(* Logix 5000 project; controller PLC_MCC1300_75F1 vendor 1 type 14 code 166 rev 32.11; software revision 32.04; part 18 of 83 *)
(* tags used below, declared in another part *)
   GP_OB_InitializeMain : GP_OB_Initialize;
   M302SpeedUp : MAC_SpeedUp;
   M310_M4_DR_B1 : AXIS_CIP_DRIVE;
   M310B : MAC_Conveyor;
   M310B_ALM : MAC_Conveyor_ALM;
   M310B_Data : UDT_Convoy_SL;
   M310B_HMR : MAC_Conveyor_HMR;
   M310B_HMW : MAC_Conveyor_HMW;
   M310B_M1_DR_IN_MAJ : MOTION_INSTRUCTION;
   M310B_M1_DR_IN_MAR : MOTION_INSTRUCTION;
   M310B_M1_DR_IN_MAS : MOTION_INSTRUCTION;
   M310B_M1_DR_IN_MRP : MOTION_INSTRUCTION;
   M310B_M1_DR_MAFR : MOTION_INSTRUCTION;
   M310B_M1_DR_MDR : MOTION_INSTRUCTION;
   M310B_M1_DR_MSF : MOTION_INSTRUCTION;
   M310B_M1_DR_MSO : MOTION_INSTRUCTION;
   M310B_M1_DR_OUT_MAJ : MOTION_INSTRUCTION;
   M310B_M1_DR_OUT_MAM : MOTION_INSTRUCTION;
   M310B_M1_DR_OUT_MAR : MOTION_INSTRUCTION;
   M310B_M1_DR_OUT_MCD : MOTION_INSTRUCTION;
   M310B_M1_DR_OUT_MRP : MOTION_INSTRUCTION;
   M310B_SpaceConv_Utilities : SpaceConv_Utilities;
   M310B_xOS_PosReq : BOOL;
   M311 : MAC_Conveyor;
   TMP_d : DINT;
   TMP_dDirection : DINT;
   TMP_r : REAL;
   TMP_rAcc : REAL;
   TMP_rDec : REAL;
   TMP_rSpeed : REAL;
   TMP_rTarget_M1 : REAL;
   TMP_xForwardCommadnForCleaningZone : BOOL;
   TMP_xPositioning : BOOL;
   TMP_xPositioning_M1 : BOOL;
   TMP_xPositioning_M2 : BOOL;
   TMP_xPowerSaving : BOOL;
   TMP_xReverse : BOOL;
   TMP_xReverse_M1 : BOOL;
   TMP_xReverse_M2 : BOOL;
   TMP_xRun : BOOL;
   TMP_xRun_M1 : BOOL;
   TMP_xRun_M2 : BOOL;
   xAlwaysOFF : BOOL;
   xAlwaysON : BOOL;
   xDebugOFF : BOOL;
   Z300_Conveyor : UDT_StandConv[29];
   Z300_Conveyor_Conf : UDT_Conveyor_Config[29];
   Z300_Conveyor_HMW : MAC_Conveyor_ZC_HMW[29];
   Z300_Conveyor_IN_MOTION : MAC_Conveyor_ZC_IN_MOTION[29];
   Z301_HMR : MAC_Zone_ML_HMR;
   Z401 : MAC_Zone;
   Z401_HMW : MAC_Zone_HMW;
(* CommandLogic, continued *)

ROUTINE M307EM1_Conveyor_Output   (* ladder *)
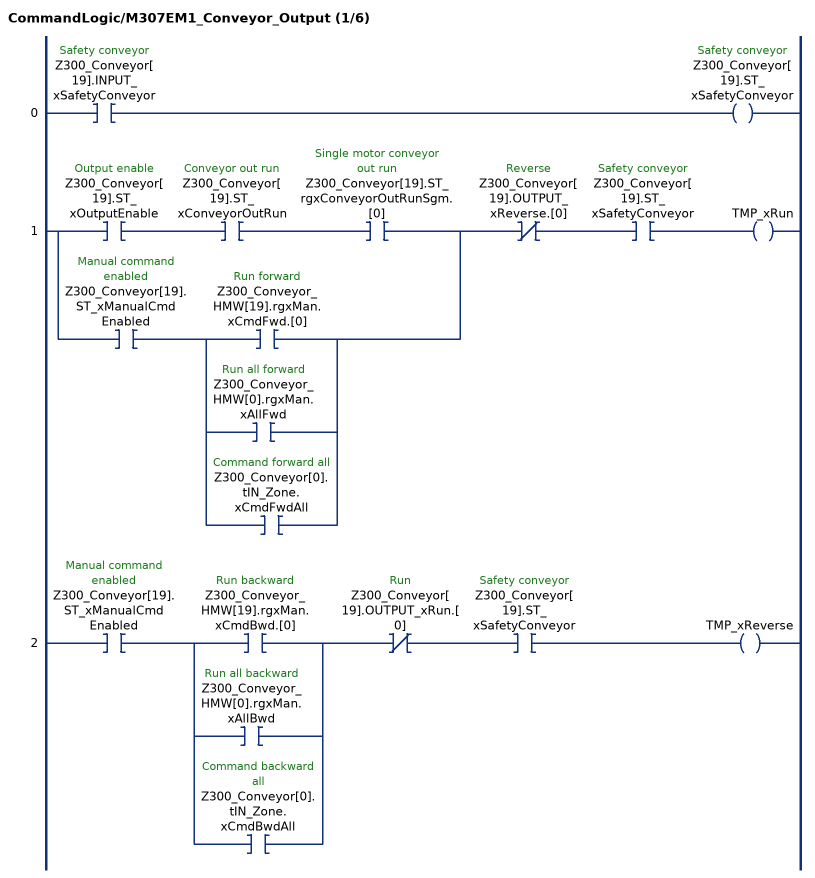
   0: XIC(Z300_Conveyor[19].INPUT_xSafetyConveyor)OTE(Z300_Conveyor[19].ST_xSafetyConveyor);
   1: [XIC(Z300_Conveyor[19].ST_xOutputEnable) XIC(Z300_Conveyor[19].ST_xConveyorOutRun) XIC(Z300_Conveyor[19].ST_rgxConveyorOutRunSgm.[0]) ,XIC(Z300_Conveyor[19].ST_xManualCmdEnabled) [XIC(Z300_Conveyor_HMW[19].rgxMan.xCmdFwd.[0]) ,XIC(Z300_Conveyor_HMW[0].rgxMan.xAllFwd) ,XIC(Z300_Conveyor[0].tIN_Zone.xCmdFwdAll) ] ]XIO(Z300_Conveyor[19].OUTPUT_xReverse.[0])XIC(Z300_Conveyor[19].ST_xSafetyConveyor)OTE(TMP_xRun);
   2: XIC(Z300_Conveyor[19].ST_xManualCmdEnabled)[XIC(Z300_Conveyor_HMW[19].rgxMan.xCmdBwd.[0]) ,XIC(Z300_Conveyor_HMW[0].rgxMan.xAllBwd) ,XIC(Z300_Conveyor[0].tIN_Zone.xCmdBwdAll) ]XIO(Z300_Conveyor[19].OUTPUT_xRun.[0])XIC(Z300_Conveyor[19].ST_xSafetyConveyor)OTE(TMP_xReverse);
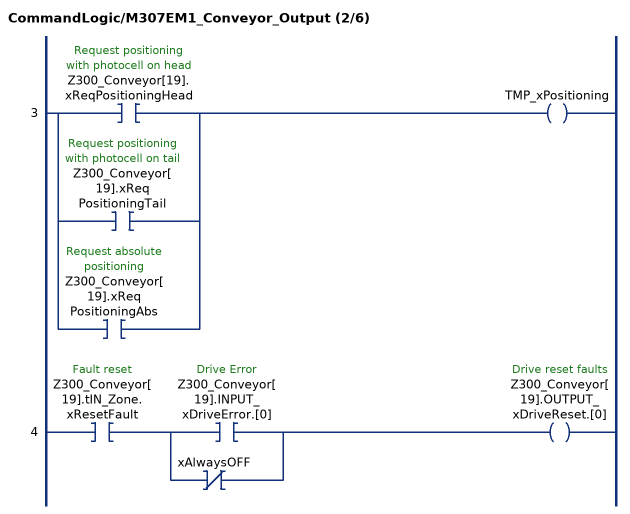
   3: [XIC(Z300_Conveyor[19].xReqPositioningHead) ,XIC(Z300_Conveyor[19].xReqPositioningTail) ,XIC(Z300_Conveyor[19].xReqPositioningAbs) ]OTE(TMP_xPositioning);
   4: XIC(Z300_Conveyor[19].tIN_Zone.xResetFault)[XIC(Z300_Conveyor[19].INPUT_xDriveError.[0]) ,XIO(xAlwaysOFF) ]OTE(Z300_Conveyor[19].OUTPUT_xDriveReset.[0]);
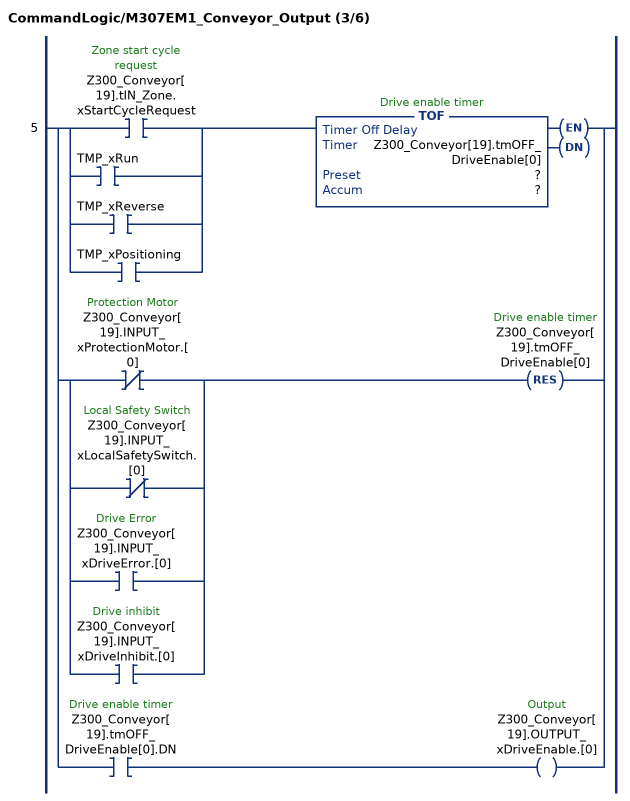
   5: [[XIC(Z300_Conveyor[19].tIN_Zone.xStartCycleRequest) ,XIC(TMP_xRun) ,XIC(TMP_xReverse) ,XIC(TMP_xPositioning) ] TOF(Z300_Conveyor[19].tmOFF_DriveEnable[0],?,?) ,[XIO(Z300_Conveyor[19].INPUT_xProtectionMotor.[0]) ,XIO(Z300_Conveyor[19].INPUT_xLocalSafetySwitch.[0]) ,XIC(Z300_Conveyor[19].INPUT_xDriveError.[0]) ,XIC(Z300_Conveyor[19].INPUT_xDriveInhibit.[0]) ] RES(Z300_Conveyor[19].tmOFF_DriveEnable[0]) ,XIC(Z300_Conveyor[19].tmOFF_DriveEnable[0].DN) OTE(Z300_Conveyor[19].OUTPUT_xDriveEnable.[0]) ];
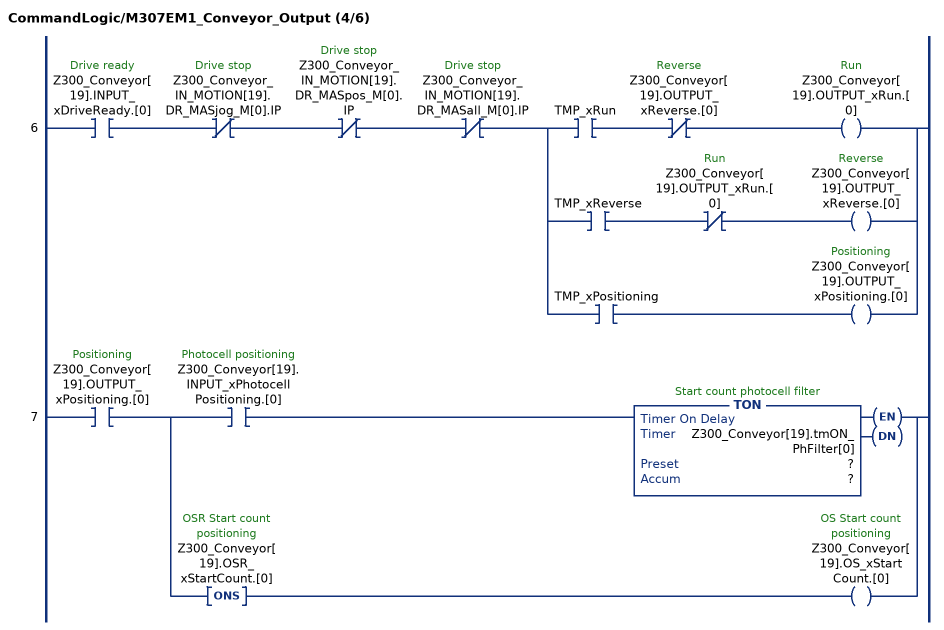
   6: XIC(Z300_Conveyor[19].INPUT_xDriveReady.[0])XIO(Z300_Conveyor_IN_MOTION[19].DR_MASjog_M[0].IP)XIO(Z300_Conveyor_IN_MOTION[19].DR_MASpos_M[0].IP)XIO(Z300_Conveyor_IN_MOTION[19].DR_MASall_M[0].IP)[XIC(TMP_xRun) XIO(Z300_Conveyor[19].OUTPUT_xReverse.[0]) OTE(Z300_Conveyor[19].OUTPUT_xRun.[0]) ,XIC(TMP_xReverse) XIO(Z300_Conveyor[19].OUTPUT_xRun.[0]) OTE(Z300_Conveyor[19].OUTPUT_xReverse.[0]) ,XIC(TMP_xPositioning) OTE(Z300_Conveyor[19].OUTPUT_xPositioning.[0]) ];
   7: XIC(Z300_Conveyor[19].OUTPUT_xPositioning.[0])[XIC(Z300_Conveyor[19].INPUT_xPhotocellPositioning.[0]) TON(Z300_Conveyor[19].tmON_PhFilter[0],?,?) ,ONS(Z300_Conveyor[19].OSR_xStartCount.[0]) OTE(Z300_Conveyor[19].OS_xStartCount.[0]) ];
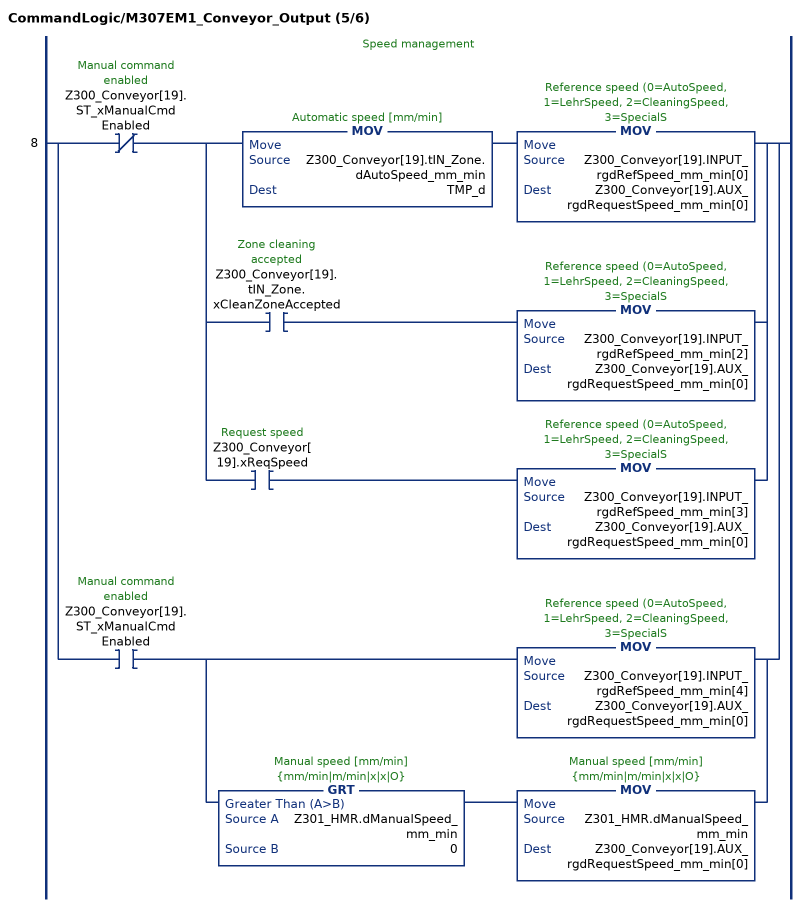
   // Speed management
   8: [XIO(Z300_Conveyor[19].ST_xManualCmdEnabled) [MOV(Z300_Conveyor[19].tIN_Zone.dAutoSpeed_mm_min,TMP_d) MOV(Z300_Conveyor[19].INPUT_rgdRefSpeed_mm_min[0],Z300_Conveyor[19].AUX_rgdRequestSpeed_mm_min[0]) ,XIC(Z300_Conveyor[19].tIN_Zone.xCleanZoneAccepted) MOV(Z300_Conveyor[19].INPUT_rgdRefSpeed_mm_min[2],Z300_Conveyor[19].AUX_rgdRequestSpeed_mm_min[0]) ,XIC(Z300_Conveyor[19].xReqSpeed) MOV(Z300_Conveyor[19].INPUT_rgdRefSpeed_mm_min[3],Z300_Conveyor[19].AUX_rgdRequestSpeed_mm_min[0]) ] ,XIC(Z300_Conveyor[19].ST_xManualCmdEnabled) [MOV(Z300_Conveyor[19].INPUT_rgdRefSpeed_mm_min[4],Z300_Conveyor[19].AUX_rgdRequestSpeed_mm_min[0]) ,GRT(Z301_HMR.dManualSpeed_mm_min,0) MOV(Z301_HMR.dManualSpeed_mm_min,Z300_Conveyor[19].AUX_rgdRequestSpeed_mm_min[0]) ] ];
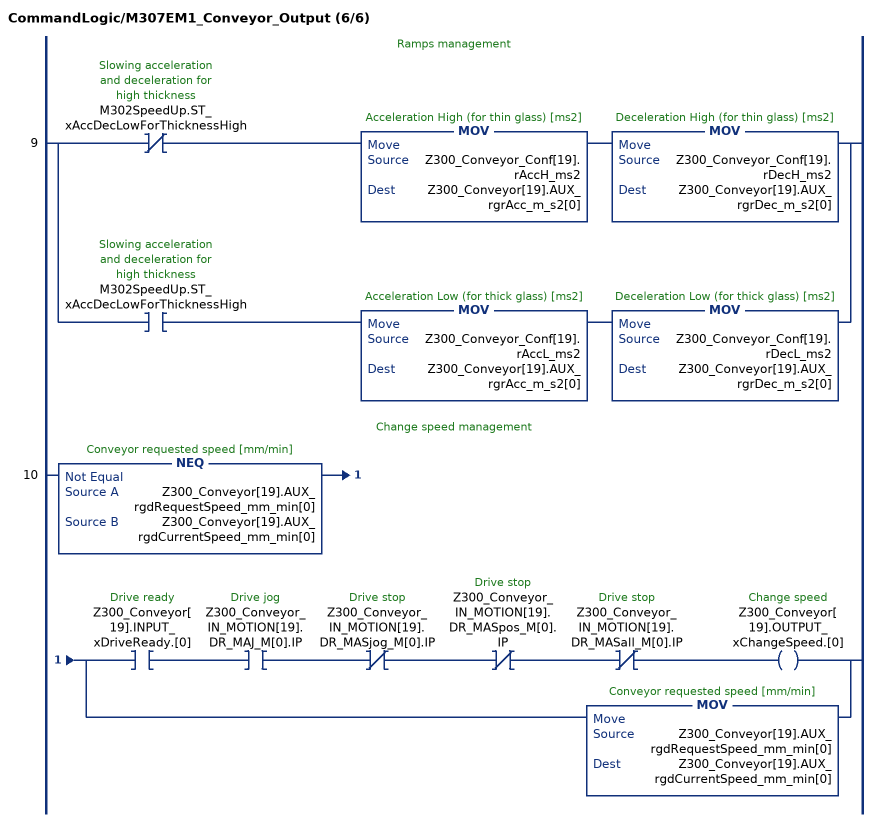
   // Ramps management
   9: [XIO(M302SpeedUp.ST_xAccDecLowForThicknessHigh) MOV(Z300_Conveyor_Conf[19].rAccH_ms2,Z300_Conveyor[19].AUX_rgrAcc_m_s2[0]) MOV(Z300_Conveyor_Conf[19].rDecH_ms2,Z300_Conveyor[19].AUX_rgrDec_m_s2[0]) ,XIC(M302SpeedUp.ST_xAccDecLowForThicknessHigh) MOV(Z300_Conveyor_Conf[19].rAccL_ms2,Z300_Conveyor[19].AUX_rgrAcc_m_s2[0]) MOV(Z300_Conveyor_Conf[19].rDecL_ms2,Z300_Conveyor[19].AUX_rgrDec_m_s2[0]) ];
   // Change speed management
   10: NEQ(Z300_Conveyor[19].AUX_rgdRequestSpeed_mm_min[0],Z300_Conveyor[19].AUX_rgdCurrentSpeed_mm_min[0])[XIC(Z300_Conveyor[19].INPUT_xDriveReady.[0]) XIC(Z300_Conveyor_IN_MOTION[19].DR_MAJ_M[0].IP) XIO(Z300_Conveyor_IN_MOTION[19].DR_MASjog_M[0].IP) XIO(Z300_Conveyor_IN_MOTION[19].DR_MASpos_M[0].IP) XIO(Z300_Conveyor_IN_MOTION[19].DR_MASall_M[0].IP) OTE(Z300_Conveyor[19].OUTPUT_xChangeSpeed.[0]) ,MOV(Z300_Conveyor[19].AUX_rgdRequestSpeed_mm_min[0],Z300_Conveyor[19].AUX_rgdCurrentSpeed_mm_min[0]) ];
END_ROUTINE

ROUTINE M307FM1_Conveyor_Output   (* ladder *)
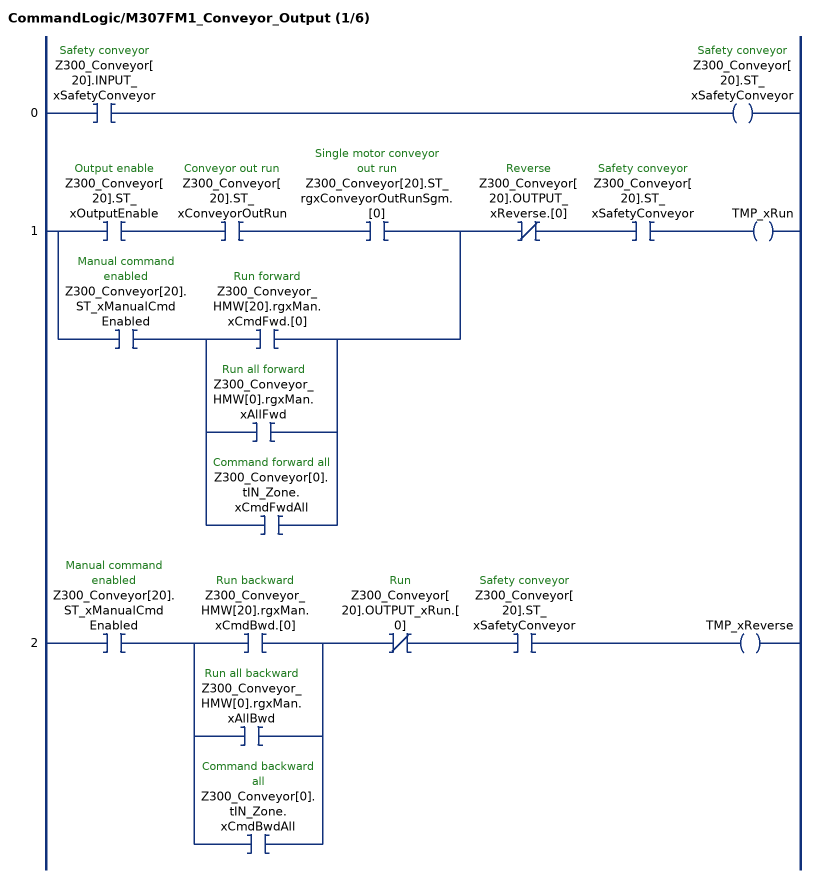
   0: XIC(Z300_Conveyor[20].INPUT_xSafetyConveyor)OTE(Z300_Conveyor[20].ST_xSafetyConveyor);
   1: [XIC(Z300_Conveyor[20].ST_xOutputEnable) XIC(Z300_Conveyor[20].ST_xConveyorOutRun) XIC(Z300_Conveyor[20].ST_rgxConveyorOutRunSgm.[0]) ,XIC(Z300_Conveyor[20].ST_xManualCmdEnabled) [XIC(Z300_Conveyor_HMW[20].rgxMan.xCmdFwd.[0]) ,XIC(Z300_Conveyor_HMW[0].rgxMan.xAllFwd) ,XIC(Z300_Conveyor[0].tIN_Zone.xCmdFwdAll) ] ]XIO(Z300_Conveyor[20].OUTPUT_xReverse.[0])XIC(Z300_Conveyor[20].ST_xSafetyConveyor)OTE(TMP_xRun);
   2: XIC(Z300_Conveyor[20].ST_xManualCmdEnabled)[XIC(Z300_Conveyor_HMW[20].rgxMan.xCmdBwd.[0]) ,XIC(Z300_Conveyor_HMW[0].rgxMan.xAllBwd) ,XIC(Z300_Conveyor[0].tIN_Zone.xCmdBwdAll) ]XIO(Z300_Conveyor[20].OUTPUT_xRun.[0])XIC(Z300_Conveyor[20].ST_xSafetyConveyor)OTE(TMP_xReverse);
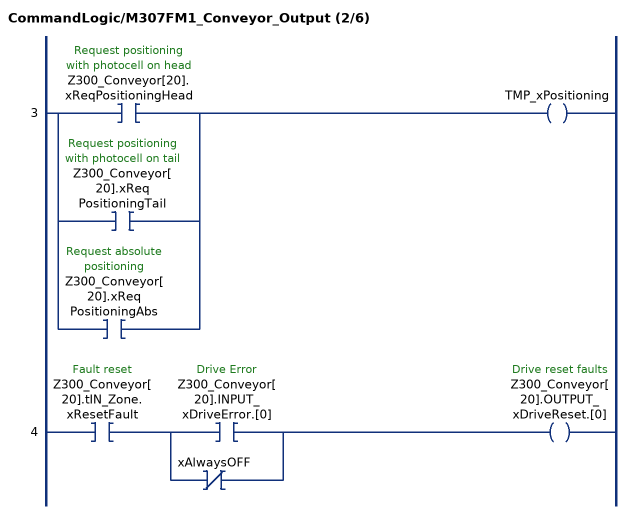
   3: [XIC(Z300_Conveyor[20].xReqPositioningHead) ,XIC(Z300_Conveyor[20].xReqPositioningTail) ,XIC(Z300_Conveyor[20].xReqPositioningAbs) ]OTE(TMP_xPositioning);
   4: XIC(Z300_Conveyor[20].tIN_Zone.xResetFault)[XIC(Z300_Conveyor[20].INPUT_xDriveError.[0]) ,XIO(xAlwaysOFF) ]OTE(Z300_Conveyor[20].OUTPUT_xDriveReset.[0]);
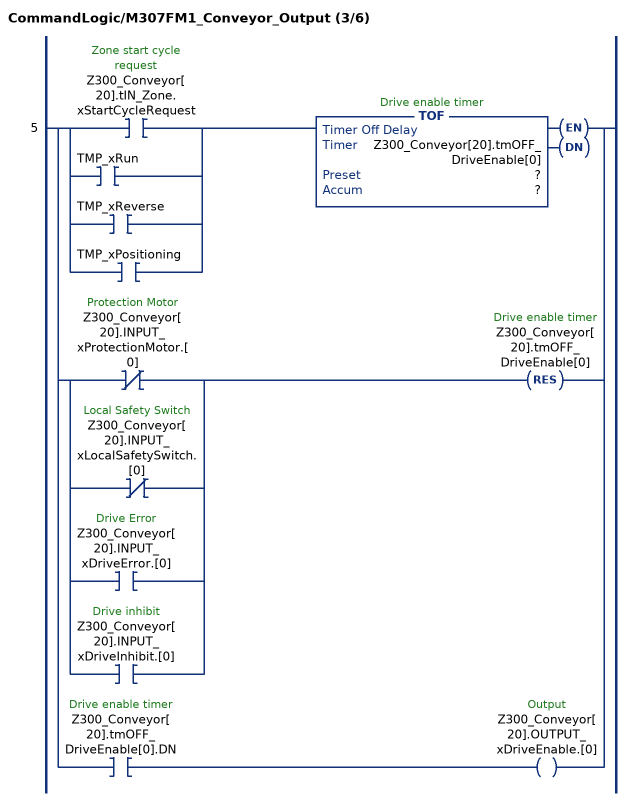
   5: [[XIC(Z300_Conveyor[20].tIN_Zone.xStartCycleRequest) ,XIC(TMP_xRun) ,XIC(TMP_xReverse) ,XIC(TMP_xPositioning) ] TOF(Z300_Conveyor[20].tmOFF_DriveEnable[0],?,?) ,[XIO(Z300_Conveyor[20].INPUT_xProtectionMotor.[0]) ,XIO(Z300_Conveyor[20].INPUT_xLocalSafetySwitch.[0]) ,XIC(Z300_Conveyor[20].INPUT_xDriveError.[0]) ,XIC(Z300_Conveyor[20].INPUT_xDriveInhibit.[0]) ] RES(Z300_Conveyor[20].tmOFF_DriveEnable[0]) ,XIC(Z300_Conveyor[20].tmOFF_DriveEnable[0].DN) OTE(Z300_Conveyor[20].OUTPUT_xDriveEnable.[0]) ];
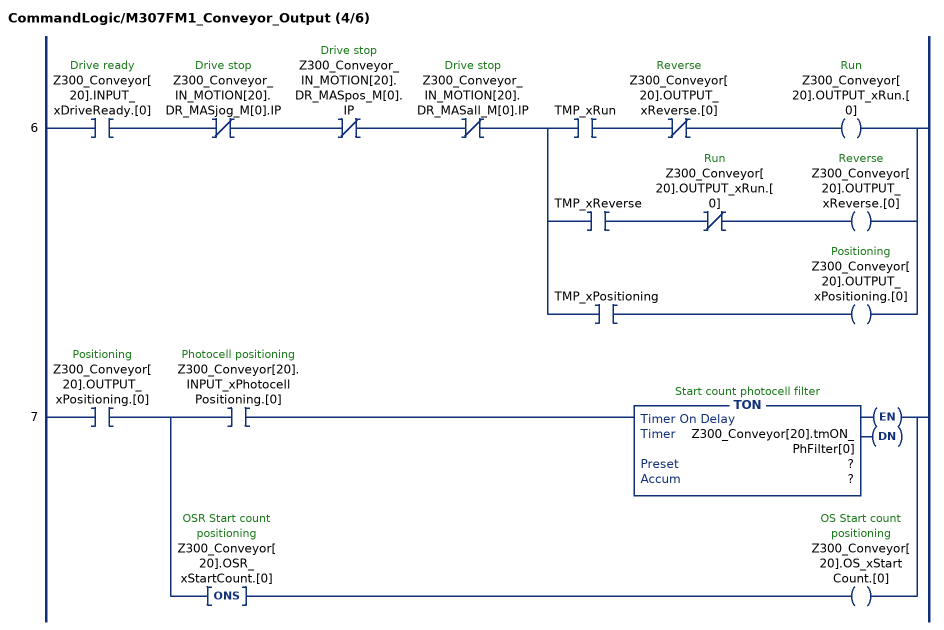
   6: XIC(Z300_Conveyor[20].INPUT_xDriveReady.[0])XIO(Z300_Conveyor_IN_MOTION[20].DR_MASjog_M[0].IP)XIO(Z300_Conveyor_IN_MOTION[20].DR_MASpos_M[0].IP)XIO(Z300_Conveyor_IN_MOTION[20].DR_MASall_M[0].IP)[XIC(TMP_xRun) XIO(Z300_Conveyor[20].OUTPUT_xReverse.[0]) OTE(Z300_Conveyor[20].OUTPUT_xRun.[0]) ,XIC(TMP_xReverse) XIO(Z300_Conveyor[20].OUTPUT_xRun.[0]) OTE(Z300_Conveyor[20].OUTPUT_xReverse.[0]) ,XIC(TMP_xPositioning) OTE(Z300_Conveyor[20].OUTPUT_xPositioning.[0]) ];
   7: XIC(Z300_Conveyor[20].OUTPUT_xPositioning.[0])[XIC(Z300_Conveyor[20].INPUT_xPhotocellPositioning.[0]) TON(Z300_Conveyor[20].tmON_PhFilter[0],?,?) ,ONS(Z300_Conveyor[20].OSR_xStartCount.[0]) OTE(Z300_Conveyor[20].OS_xStartCount.[0]) ];
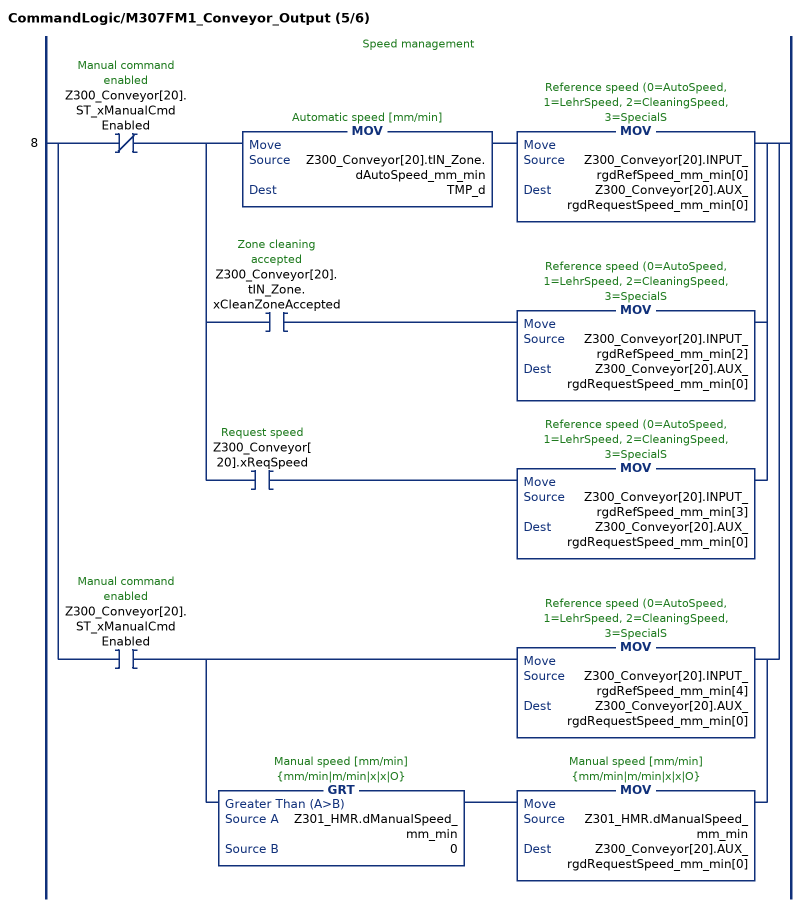
   // Speed management
   8: [XIO(Z300_Conveyor[20].ST_xManualCmdEnabled) [MOV(Z300_Conveyor[20].tIN_Zone.dAutoSpeed_mm_min,TMP_d) MOV(Z300_Conveyor[20].INPUT_rgdRefSpeed_mm_min[0],Z300_Conveyor[20].AUX_rgdRequestSpeed_mm_min[0]) ,XIC(Z300_Conveyor[20].tIN_Zone.xCleanZoneAccepted) MOV(Z300_Conveyor[20].INPUT_rgdRefSpeed_mm_min[2],Z300_Conveyor[20].AUX_rgdRequestSpeed_mm_min[0]) ,XIC(Z300_Conveyor[20].xReqSpeed) MOV(Z300_Conveyor[20].INPUT_rgdRefSpeed_mm_min[3],Z300_Conveyor[20].AUX_rgdRequestSpeed_mm_min[0]) ] ,XIC(Z300_Conveyor[20].ST_xManualCmdEnabled) [MOV(Z300_Conveyor[20].INPUT_rgdRefSpeed_mm_min[4],Z300_Conveyor[20].AUX_rgdRequestSpeed_mm_min[0]) ,GRT(Z301_HMR.dManualSpeed_mm_min,0) MOV(Z301_HMR.dManualSpeed_mm_min,Z300_Conveyor[20].AUX_rgdRequestSpeed_mm_min[0]) ] ];